   "3#冲渣泵电动阀开" AT %Q22.5 : Bool;
   "3#冲渣泵电动阀关" AT %Q22.6 : Bool;
   "3#冲渣泵排气电磁阀" AT %Q22.7 : Bool;
   "2#冲渣泵引水电磁阀" AT %Q23.0 : Bool;
   "2#冲渣泵电动阀开" AT %Q23.1 : Bool;
   "2#冲渣泵电动阀关" AT %Q23.2 : Bool;
   "2#冲渣泵排气电磁阀" AT %Q23.3 : Bool;
   "1#冲渣泵引水电磁阀" AT %Q23.4 : Bool;
   "1#冲渣泵电动阀开" AT %Q23.5 : Bool;
   "1#冲渣泵电动阀关" AT %Q23.6 : Bool;
   "1#冲渣泵排气电磁阀" AT %Q23.7 : Bool;
   "1#冲渣泵管道压力" AT %IW368 : Int;
   "2#冲渣泵管道压力" AT %IW370 : Int;
   "3#冲渣泵管道压力" AT %IW372 : Int;
   "4#冲渣泵管道压力" AT %IW374 : Int;
   "5#冲渣泵管道压力" AT %IW376 : Int;
   "6#冲渣泵管道压力" AT %IW378 : Int;
   "7#冲渣泵管道压力" AT %IW380 : Int;
   "8#冲渣泵管道压力" AT %IW382 : Int;
   "1#冲渣阀门开度" AT %IW384 : Int;
   "2#冲渣阀门开度" AT %IW386 : Int;
   "3#冲渣阀门开度" AT %IW388 : Int;
   "4#冲渣阀门开度" AT %IW390 : Int;
   "5#冲渣阀门开度" AT %IW392 : Int;
   "6#冲渣阀门开度" AT %IW394 : Int;
   "7#冲渣阀门开度" AT %IW396 : Int;
   "8#冲渣阀门开度" AT %IW398 : Int;
   "1#冲渣泵阀门开度给定" AT %QW320 : Int;
   "2#冲渣泵阀门开度给定" AT %QW322 : Int;
   "3#冲渣泵阀门开度给定" AT %QW324 : Int;
   "4#冲渣泵阀门开度给定" AT %QW326 : Int;
   "5#冲渣泵阀门开度给定" AT %QW328 : Int;
   "6#冲渣泵阀门开度给定" AT %QW330 : Int;
   "7#冲渣泵阀门开度给定" AT %QW332 : Int;
   "8#冲渣泵阀门开度给定" AT %QW334 : Int;
   "窑冷却泵运行" AT %I23.6 : Bool;
   "窑冷却泵故障" AT %I23.7 : Bool;
   "窑冷却泵驱动" AT %Q4.7 : Bool;
   "5#净环热水泵驱动" AT %Q5.0 : Bool;
   "Q5_1" AT %Q5.1 : Bool;
   "Q5_2" AT %Q5.2 : Bool;
   "Q5_3" AT %Q5.3 : Bool;
   "Q5_4" AT %Q5.4 : Bool;
   "Q5_5" AT %Q5.5 : Bool;
   "Q5_6" AT %Q5.6 : Bool;
   "Q5_7" AT %Q5.7 : Bool;
   "Q6_0" AT %Q6.0 : Bool;
   "Q6_1" AT %Q6.1 : Bool;
   "Q6_2" AT %Q6.2 : Bool;
   "Q6_3" AT %Q6.3 : Bool;
   "Q6_4" AT %Q6.4 : Bool;
   "Q6_5" AT %Q6.5 : Bool;
   "Q6_6" AT %Q6.6 : Bool;
   "Q6_7" AT %Q6.7 : Bool;
   "Q7_0" AT %Q7.0 : Bool;
   "Q7_1" AT %Q7.1 : Bool;
   "Q7_2" AT %Q7.2 : Bool;
   "Q7_3" AT %Q7.3 : Bool;
   "Q7_4" AT %Q7.4 : Bool;
   "Q7_5" AT %Q7.5 : Bool;
   "Q7_6" AT %Q7.6 : Bool;
   "Q7_7" AT %Q7.7 : Bool;
   "I32_6" AT %I32.6 : Bool;
   "I32_7" AT %I32.7 : Bool;
   "窑冷却泵电动蝶阀备妥" AT %I33.0 : Bool;
   "窑冷却泵电动蝶阀运行" AT %I33.1 : Bool;
   "窑冷却泵电动蝶阀故障" AT %I33.2 : Bool;
   "窑冷却泵电动蝶阀开到位" AT %I33.3 : Bool;
   "窑冷却泵电动蝶阀关到位" AT %I33.4 : Bool;
   "I33_5" AT %I33.5 : Bool;
   "I33_6" AT %I33.6 : Bool;
   "I33_7" AT %I33.7 : Bool;
   "I34_0" AT %I34.0 : Bool;
   "I34_1" AT %I34.1 : Bool;
   "I34_2" AT %I34.2 : Bool;
   "I34_3" AT %I34.3 : Bool;
   "I34_4" AT %I34.4 : Bool;
   "I34_5" AT %I34.5 : Bool;
   "I34_6" AT %I34.6 : Bool;
   "I34_7" AT %I34.7 : Bool;
   "I35_0" AT %I35.0 : Bool;
   "I35_1" AT %I35.1 : Bool;
   "I35_2" AT %I35.2 : Bool;
   "I35_3" AT %I35.3 : Bool;
   "I35_4" AT %I35.4 : Bool;
   "I35_5" AT %I35.5 : Bool;
   "I35_6" AT %I35.6 : Bool;
   "I35_7" AT %I35.7 : Bool;
   "5#净环热水泵电动阀开" AT %Q14.0 : Bool;
   "5#净环热水泵电动阀关" AT %Q14.1 : Bool;
   "窑冷却泵电动阀开" AT %Q14.2 : Bool;
   "窑冷却泵电动阀关" AT %Q14.3 : Bool;
   "1#柴油泵电动阀开" AT %Q14.4 : Bool;
   "1#柴油泵电动阀关" AT %Q14.5 : Bool;
   "2#柴油泵电动阀开" AT %Q14.6 : Bool;
   "2#柴油泵电动阀关" AT %Q14.7 : Bool;
   "Q15_0" AT %Q15.0 : Bool;
   "Q15_1" AT %Q15.1 : Bool;
   "Q15_2" AT %Q15.2 : Bool;
   "Q15_3" AT %Q15.3 : Bool;
   "Q15_4" AT %Q15.4 : Bool;
   "Q15_5" AT %Q15.5 : Bool;
   "Q15_6" AT %Q15.6 : Bool;
   "Q15_7" AT %Q15.7 : Bool;
   "PIW322" AT %IW322 : Int;
   "PIW324" AT %IW324 : Int;
   "PIW326" AT %IW326 : Int;
   "PIW328" AT %IW328 : Int;
   "PIW330" AT %IW330 : Int;
   "PIW332" AT %IW332 : Int;
   "PIW334" AT %IW334 : Int;
   "PQW290" AT %QW290 : Int;
   "PQW292" AT %QW292 : Int;
   "PQW294" AT %QW294 : Int;
   "PQW296" AT %QW296 : Int;
   "PQW298" AT %QW298 : Int;
   "PQW300" AT %QW300 : Int;
   "PQW302" AT %QW302 : Int;
   "I41_0" AT %I41.0 : Bool;
   "I41_1" AT %I41.1 : Bool;
   "I41_2" AT %I41.2 : Bool;
   "I41_3" AT %I41.3 : Bool;
   "I41_4" AT %I41.4 : Bool;
   "I41_5" AT %I41.5 : Bool;
   "I41_6" AT %I41.6 : Bool;
   "I41_7" AT %I41.7 : Bool;
   "I42_0" AT %I42.0 : Bool;
   "I42_1" AT %I42.1 : Bool;
   "I42_2" AT %I42.2 : Bool;
   "I42_3" AT %I42.3 : Bool;
   "I42_4" AT %I42.4 : Bool;
   "I42_5" AT %I42.5 : Bool;
   "I42_6" AT %I42.6 : Bool;
   "I42_7" AT %I42.7 : Bool;
   "I43_0" AT %I43.0 : Bool;
   "I43_1" AT %I43.1 : Bool;
   "I43_2" AT %I43.2 : Bool;
   "I43_3" AT %I43.3 : Bool;
   "I43_4" AT %I43.4 : Bool;
   "I43_5" AT %I43.5 : Bool;
   "I43_6" AT %I43.6 : Bool;
   "I43_7" AT %I43.7 : Bool;
   "I49_0" AT %I49.0 : Bool;
   "I49_1" AT %I49.1 : Bool;
   "I49_2" AT %I49.2 : Bool;
   "I49_3" AT %I49.3 : Bool;
   "I49_4" AT %I49.4 : Bool;
   "I49_5" AT %I49.5 : Bool;
   "I49_6" AT %I49.6 : Bool;
   "I49_7" AT %I49.7 : Bool;
   "I50_0" AT %I50.0 : Bool;
   "I50_1" AT %I50.1 : Bool;
   "I50_2" AT %I50.2 : Bool;
   "I50_3" AT %I50.3 : Bool;
   "I50_4" AT %I50.4 : Bool;
   "I50_5" AT %I50.5 : Bool;
   "I50_6" AT %I50.6 : Bool;
   "I50_7" AT %I50.7 : Bool;
   "I51_0" AT %I51.0 : Bool;
   "I51_1" AT %I51.1 : Bool;
   "I51_2" AT %I51.2 : Bool;
   "I51_3" AT %I51.3 : Bool;
   "I51_4" AT %I51.4 : Bool;
   "I51_5" AT %I51.5 : Bool;
   "I51_6" AT %I51.6 : Bool;
   "I51_7" AT %I51.7 : Bool;
   "Tag_1" AT %M1.4 : Bool;
   "Tag_2" AT %M2.0 : Bool;
   "Tag_3" AT %T40 : Timer;
   "Tag_4" AT %M2.1 : Bool;
   "Tag_5" AT %MW4 : Int;
   "Tag_6" AT %M2.2 : Bool;
   "Tag_7" AT %M2.3 : Bool;
   "Tag_8" AT %M2.4 : Bool;
   "Tag_9" AT %M2.5 : Bool;
   "Tag_10" AT %M2.6 : Bool;
   "Tag_11" AT %M2.7 : Bool;
   "Tag_12" AT %M3.0 : Bool;
   "Tag_13" AT %M3.1 : Bool;
   "Tag_14" AT %M3.2 : Bool;
   "Tag_15" AT %MD4 : Real;
   "Tag_16" AT %MD8 : Real;
   "HMI_允许电炉启动冲渣泵1" AT %M100.0 : Bool;
   "HMI_允许电炉启动冲渣泵2" AT %M100.1 : Bool;
   "HMI_允许电炉启动冲渣泵3" AT %M100.2 : Bool;
   "HMI_允许电炉启动冲渣泵4" AT %M100.3 : Bool;
   "HMI_允许电炉启动冲渣泵5" AT %M100.4 : Bool;
   "HMI_允许电炉启动冲渣泵6" AT %M100.5 : Bool;
   "HMI_允许电炉启动冲渣泵7" AT %M100.6 : Bool;
   "HMI_允许电炉启动冲渣泵8" AT %M100.7 : Bool;
   "HMI_电炉冲渣急停1" AT %M99.0 : Bool;
   "HMI_电炉冲渣急停2" AT %M99.1 : Bool;
   "Tag_17" AT %M11.1 : Bool;
END_VAR

DATA_BLOCK "AI"   // DB2
{ S7_Optimized_Access := 'FALSE' }
VERSION : 0.1
   VAR
      "1#炉体水泵管道压力" : Real;
      "2#炉体水泵管道压力" : Real;
      "3#炉体水泵管道压力" : Real;
      "1#电极水泵管道压力" : Real;
      "2#电极水泵管道压力" : Real;
      "3#电极水泵管道压力" : Real;
      "4#电极水泵管道压力" : Real;
      "1#柴油泵管道压力" : Real;
      "2#柴油泵管道压力" : Real;
      "1#炉体水阀门开度" : Real;
      "2#炉体水阀门开度" : Real;
      "3#炉体水阀门开度" : Real;
      "1#电极水阀门开度" : Real;
      "2#电极水阀门开度" : Real;
      "3#电极水阀门开度" : Real;
      "4#电极水阀门开度" : Real;
      "2#柴油泵阀门开度" : Real;
      "1#净环热水管道压力" : Real;
      "2#净环热水管道压力" : Real;
      "3#净环热水管道压力" : Real;
      "4#净环热水管道压力" : Real;
      "5#净环热水管道压力" : Real;
      "6#净环热水管道压力" : Real;
      "1#净环热水阀门开度" : Real;
      "2#净环热水阀门开度" : Real;
      "3#净环热水阀门开度" : Real;
      "4#净环热水阀门开度" : Real;
      "5#净环热水阀门开度" : Real;
      "6#净环热水阀门开度" : Real;
      "1#外围补水阀门开度" : Real;
      "2#外围补水阀门开度" : Real;
      "1#水池液位" : Real;
      "2#水池液位" : Real;
      PIW322 : Real;
      PIW324 : Real;
      PIW326 : Real;
      PIW328 : Real;
      PIW330 : Real;
      PIW332 : Real;
      PIW334 : Real;
      "1#冲渣热水泵管道压力" : Real;
      "2#冲渣热水泵管道压力" : Real;
      "3#冲渣热水泵管道压力" : Real;
      "4#冲渣热水泵管道压力" : Real;
      "5#冲渣热水泵管道压力" : Real;
      "6#冲渣热水泵管道压力" : Real;
      "7#冲渣热水泵管道压力" : Real;
      "8#冲渣热水泵管道压力" : Real;
      "1#冲渣热水阀门开度" : Real;
      "2#冲渣热水阀门开度" : Real;
      "3#冲渣热水阀门开度" : Real;
      "4#冲渣热水阀门开度" : Real;
      "5#冲渣热水阀门开度" : Real;
      "6#冲渣热水阀门开度" : Real;
      "7#冲渣热水阀门开度" : Real;
      "8#冲渣热水阀门开度" : Real;
      "1#冲渣泵管道压力" : Real;
      "2#冲渣泵管道压力" : Real;
      "3#冲渣泵管道压力" : Real;
      "4#冲渣泵管道压力" : Real;
      "5#冲渣泵管道压力" : Real;
      "6#冲渣泵管道压力" : Real;
      "7#冲渣泵管道压力" : Real;
      "8#冲渣泵管道压力" : Real;
      "1#冲渣阀门开度" : Real;
      "2#冲渣阀门开度" : Real;
      "3#冲渣阀门开度" : Real;
      "4#冲渣阀门开度" : Real;
      "5#冲渣阀门开度" : Real;
      "6#冲渣阀门开度" : Real;
      "7#冲渣阀门开度" : Real;
      "8#冲渣阀门开度" : Real;
      Static1 : Real;
      Static2 : Real;
      Static3 : Real;
      Static4 : Real;
      Static5 : Real;
      Static6 : Real;
      Static7 : Real;
      Static8 : Real;
      Static9 : Real;
      Static10 : Real;
      Static11 : Real;
      Static12 : Real;
      Static13 : Real;
      Static14 : Real;
      Static15 : Real;
      Static16 : Real;
      Static17 : Real;
      Static18 : Real;
      Static19 : Real;
      Static20 : Real;
      Static21 : Real;
      Static22 : Real;
      Static23 : Real;
      Static24 : Real;
      Static25 : Real;
      Static26 : Real;
      Static27 : Real;
      Static28 : Real;
      Static29 : Real;
      Static30 : Real;
      Static31 : Real;
      Static32 : Real;
      Static33 : Real;
      Static34 : Real;
      Static35 : Real;
      Static36 : Real;
      Static37 : Real;
      Static38 : Real;
      Static39 : Real;
      Static40 : Real;
      Static41 : Real;
      Static42 : Real;
      Static43 : Real;
      Static44 : Real;
      Static45 : Real;
      Static46 : Real;
      Static47 : Real;
      Static48 : Real;
      Static49 : Real;
      Static50 : Real;
      Static51 : Real;
      Static52 : Real;
      Static53 : Real;
      Static54 : Real;
      Static55 : Real;
      Static56 : Real;
      Static57 : Real;
      Static58 : Real;
      Static59 : Real;
      Static60 : Real;
      Static61 : Real;
      Static62 : Real;
      Static63 : Real;
      Static64 : Real;
      Static65 : Real;
      Static66 : Real;
      Static67 : Real;
      Static68 : Real;
      Static69 : Real;
      Static70 : Real;
      Static71 : Real;
      Static72 : Real;
      Static73 : Real;
      Static74 : Real;
      Static75 : Real;
      Static76 : Real;
      Static77 : Real;
      Static78 : Real;
      Static79 : Real;
      Static80 : Real;
      Static81 : Real;
      Static82 : Real;
      Static83 : Real;
      Static84 : Real;
      Static85 : Real;
      Static86 : Real;
      Static87 : Real;
      Static88 : Real;
      Static89 : Real;
      Static90 : Real;
      Static91 : Real;
      Static92 : Real;
      Static93 : Real;
      Static94 : Real;
      Static95 : Real;
      Static96 : Real;
      Static97 : Real;
      Static98 : Real;
      Static99 : Real;
   END_VAR
BEGIN
END_DATA_BLOCK

DATA_BLOCK "AO"   // DB3
{ S7_Optimized_Access := 'TRUE' }
VERSION : 0.1
   VAR
      "1#循环水泵阀门开度给定" : Real := 0.0;
      "2#循环水泵阀门开度给定" : Real := 0.0;
      "3#循环水泵阀门开度给定" : Real := 0.0;
      "1#电极冷却泵阀门开度给定" : Real := 0.0;
      "2#电极冷却泵阀门开度给定" : Real := 0.0;
      "3#电极冷却泵阀门开度给定" : Real := 0.0;
      "4#电极冷却泵阀门开度给定" : Real := 0.0;
      "1#柴油泵阀门开度给定" : Real := 0.0;
      "2#柴油泵阀门开度给定" : Real := 0.0;
      "1#净环热水泵阀门开度给定" : Real := 0.0;
      "2#净环热水泵阀门开度给定" : Real := 0.0;
      "3#净环热水泵阀门开度给定" : Real := 0.0;
      "4#净环热水泵阀门开度给定" : Real := 0.0;
      "5#净环热水泵阀门开度给定" : Real := 0.0;
      "6#净环热水泵阀门开度给定" : Real := 0.0;
      "1#外围补水阀门开度给定" : Real := 0.0;
      "2#外围补水阀门开度给定" : Real := 0.0;
      PQW290 : Real := 0.0;   // useless
      PQW292 : Real := 0.0;
      PQW294 : Real := 0.0;
      PQW296 : Real := 0.0;
      PQW298 : Real := 0.0;
      PQW300 : Real := 0.0;
      PQW302 : Real := 0.0;
      "1#冲渣热水泵阀门开度给定" : Real := 0.0;
      "2#冲渣热水泵阀门开度给定" : Real := 0.0;
      "3#冲渣热水泵阀门开度给定" : Real := 0.0;
      "4#冲渣热水泵阀门开度给定" : Real := 0.0;
      "5#冲渣热水泵阀门开度给定" : Real := 0.0;
      "6#冲渣热水泵阀门开度给定" : Real := 0.0;
      "7#冲渣热水泵阀门开度给定" : Real := 0.0;
      "8#冲渣热水泵阀门开度给定" : Real := 0.0;
      "1#冲渣泵阀门开度给定" : Real := 0.0;
      "2#冲渣泵阀门开度给定" : Real := 0.0;
      "3#冲渣泵阀门开度给定" : Real := 0.0;
      "4#冲渣泵阀门开度给定" : Real := 0.0;
      "5#冲渣泵阀门开度给定" : Real := 0.0;
      "6#冲渣泵阀门开度给定" : Real := 0.0;
      "7#冲渣泵阀门开度给定" : Real := 0.0;
      "8#冲渣泵阀门开度给定" : Real := 0.0;
      Static1 : Real := 0.0;
      Static2 : Real := 0.0;
      Static3 : Real := 0.0;
      Static4 : Real := 0.0;
      Static5 : Real := 0.0;
      Static6 : Real := 0.0;
      Static7 : Real := 0.0;
      Static8 : Real := 0.0;
      Static9 : Real := 0.0;
      Static10 : Real := 0.0;
      Static11 : Real := 0.0;
      Static12 : Real := 0.0;
      Static13 : Real := 0.0;
      Static14 : Real := 0.0;
      Static15 : Real := 0.0;
      Static16 : Real := 0.0;
      Static17 : Real := 0.0;
      Static18 : Real := 0.0;
      Static19 : Real := 0.0;
      Static20 : Real := 0.0;
      Static21 : Real := 0.0;
      Static22 : Real := 0.0;
      Static23 : Real := 0.0;
      Static24 : Real := 0.0;
      Static25 : Real := 0.0;
      Static26 : Real := 0.0;
      Static27 : Real := 0.0;
      Static28 : Real := 0.0;
      Static29 : Real := 0.0;
      Static30 : Real := 0.0;
      Static31 : Real := 0.0;
      Static32 : Real := 0.0;
      Static33 : Real := 0.0;
      Static34 : Real := 0.0;
      Static35 : Real := 0.0;
      Static36 : Real := 0.0;
      Static37 : Real := 0.0;
      Static38 : Real := 0.0;
      Static39 : Real := 0.0;
      Static40 : Real := 0.0;
      Static41 : Real := 0.0;
      Static42 : Real := 0.0;
      Static43 : Real := 0.0;
      Static44 : Real := 0.0;
      Static45 : Real := 0.0;
      Static46 : Real := 0.0;
      Static47 : Real := 0.0;
      Static48 : Real := 0.0;
      Static49 : Real := 0.0;
      Static50 : Real := 0.0;
      Static51 : Real := 0.0;
      Static52 : Real := 0.0;
      Static53 : Real := 0.0;
      Static54 : Real := 0.0;
      Static55 : Real := 0.0;
      Static56 : Real := 0.0;
      Static57 : Real := 0.0;
      Static58 : Real := 0.0;
      Static99 : Real := 0.0;
   END_VAR
BEGIN
END_DATA_BLOCK

DATA_BLOCK "TIME"   // DB4
{ S7_Optimized_Access := 'TRUE' }
VERSION : 0.1
   VAR
      T1 : IEC_TIMER;
      T2 : IEC_TIMER;
      T3 : IEC_TIMER;
      T4 : IEC_TIMER;
      T5 : IEC_TIMER;
      T6 : IEC_TIMER;
      T7 : IEC_TIMER;
      T8 : IEC_TIMER;
      T9 : IEC_TIMER;
      T10 : IEC_TIMER;
      T11 : IEC_TIMER;
      T12 : IEC_TIMER;
      T13 : IEC_TIMER;
      T14 : IEC_TIMER;
      T15 : IEC_TIMER;
      T16 : IEC_TIMER;
      T17 : IEC_TIMER;
      T18 : IEC_TIMER;
      T19 : IEC_TIMER;
      T20 : IEC_TIMER;
      T21 : IEC_TIMER;
      T22 : IEC_TIMER;
      T23 : IEC_TIMER;
      T24 : IEC_TIMER;
      T25 : IEC_TIMER;
      T26 : IEC_TIMER;
      T27 : IEC_TIMER;
      T28 : IEC_TIMER;
   END_VAR
BEGIN
END_DATA_BLOCK

DATA_BLOCK "DB15_PLC_TO_HMI"   // DB5
{ S7_Optimized_Access := 'FALSE' }
VERSION : 0.1
   VAR
      P1 : Bool;
      P2 : Bool;
      P3 : Bool;
      P4 : Bool;
      P5 : Bool;
      P6 : Bool;
      P7 : Bool;
      P8 : Bool;
      P9 : Bool;
      P10 : Bool;
      P11 : Bool;
      P12 : Bool;
      P13 : Bool;
      P14 : Bool;
      P15 : Bool;
      P16 : Bool;
      HMI_电炉冲渣急停1次数 : Int;
      HMI_电炉冲渣急停2次数 : Int;
      static1 : Int;
      static2 : Int;
      static3 : Int;
      static4 : Int;
      static5 : Int;
      static6 : Int;
      static7 : Int;
      static8 : Int;
      static9 : Int;
      static10 : Int;
      static11 : Int;
      static12 : Int;
   END_VAR
BEGIN
END_DATA_BLOCK

DATA_BLOCK "电机_冷却塔风机FB_DB"   // DB10
{ S7_Optimized_Access := 'FALSE' }
VERSION : 0.1
// stored: InstanceOfName 电机_冷却塔风机FB
"电机_冷却塔风机FB"
BEGIN
END_DATA_BLOCK

DATA_BLOCK "阀门_FB_DB"   // DB11
{ S7_Optimized_Access := 'FALSE' }
VERSION : 0.1
// stored: InstanceOfName 阀门_FB
"阀门_FB"
BEGIN
END_DATA_BLOCK

DATA_BLOCK "引水阀和排气阀FB_DB"   // DB12
{ S7_Optimized_Access := 'FALSE' }
VERSION : 0.1
// stored: InstanceOfName 引水阀和排气阀FB
"引水阀和排气阀FB"
BEGIN
END_DATA_BLOCK

DATA_BLOCK "电机_泵FB_DB"   // DB13
{ S7_Optimized_Access := 'FALSE' }
VERSION : 0.1
// stored: InstanceOfName 电机_泵FB
"电机_泵FB"
BEGIN
END_DATA_BLOCK

DATA_BLOCK "FB14_DATA_ALARM_DB"   // DB14
{ S7_Optimized_Access := 'FALSE' }
VERSION : 0.1
// stored: InstanceOfName FB14_DATA_ALARM
"FB14_DATA_ALARM"
BEGIN
END_DATA_BLOCK

DATA_BLOCK "FB15_MOTOR_AUTO-st_DB"   // DB15
{ S7_Optimized_Access := 'FALSE' }
VERSION : 0.1
// stored: InstanceOfName FB15_MOTOR_AUTO-st
"FB15_MOTOR_AUTO-st"
BEGIN
END_DATA_BLOCK

FUNCTION_BLOCK "电机_冷却塔风机FB"   // FB10, LAD
{ S7_Optimized_Access := 'FALSE' }
VERSION : 0.1
   VAR
      "1#冲渣水池冷却塔风机" : "电机_冷却塔风机";
      "2#冲渣水池冷却塔风机" : "电机_冷却塔风机";
      "3#冲渣水池冷却塔风机" : "电机_冷却塔风机";
      "4#冲渣水池冷却塔风机" : "电机_冷却塔风机";
      "5#冲渣水池冷却塔风机" : "电机_冷却塔风机";
      "6#冲渣水池冷却塔风机" : "电机_冷却塔风机";
      "1#净环水池冷却塔风机" : "电机_冷却塔风机";
      "2#净环水池冷却塔风机" : "电机_冷却塔风机";
      "3#净环水池冷却塔风机" : "电机_冷却塔风机";
      "4#净环水池冷却塔风机" : "电机_冷却塔风机";
      备用1 : "电机_冷却塔风机";
      备用2 : "电机_冷却塔风机";
      备用3 : "电机_冷却塔风机";
      备用4 : "电机_冷却塔风机";
      备用5 : "电机_冷却塔风机";
      备用6 : "电机_冷却塔风机";
      备用7 : "电机_冷却塔风机";
      备用8 : "电机_冷却塔风机";
      备用9 : "电机_冷却塔风机";
      备用10 : "电机_冷却塔风机";
   END_VAR
BEGIN

REGION Network 1
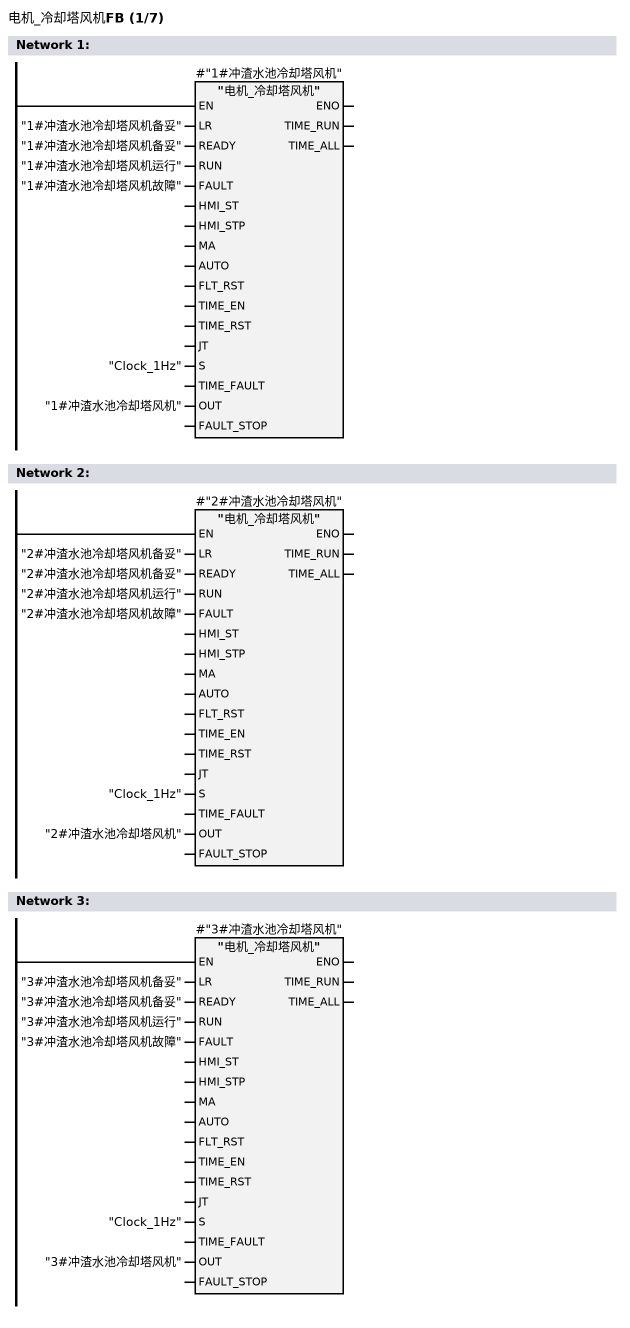
   RUNG wire#powerrail
      #"1#冲渣水池冷却塔风机"(LR := "1#冲渣水池冷却塔风机备妥", READY := "1#冲渣水池冷却塔风机备妥", RUN := "1#冲渣水池冷却塔风机运行", FAULT := "1#冲渣水池冷却塔风机故障", HMI_ST :=, HMI_STP :=, MA :=, AUTO :=, FLT_RST :=, TIME_EN :=, TIME_RST :=, JT :=, S := "Clock_1Hz", TIME_FAULT :=, OUT := "1#冲渣水池冷却塔风机", FAULT_STOP :=, TIME_RUN =>, TIME_ALL =>)
   END_RUNG
   // the same network as SCL:
   #"1#冲渣水池冷却塔风机"(LR := "1#冲渣水池冷却塔风机备妥",   // "电机_冷却塔风机"
                  READY := "1#冲渣水池冷却塔风机备妥",
                  RUN := "1#冲渣水池冷却塔风机运行",
                  FAULT := "1#冲渣水池冷却塔风机故障",
                  S := "Clock_1Hz",
                  OUT := "1#冲渣水池冷却塔风机");
END_REGION

REGION Network 2
   RUNG wire#powerrail
      #"2#冲渣水池冷却塔风机"(LR := "2#冲渣水池冷却塔风机备妥", READY := "2#冲渣水池冷却塔风机备妥", RUN := "2#冲渣水池冷却塔风机运行", FAULT := "2#冲渣水池冷却塔风机故障", HMI_ST :=, HMI_STP :=, MA :=, AUTO :=, FLT_RST :=, TIME_EN :=, TIME_RST :=, JT :=, S := "Clock_1Hz", TIME_FAULT :=, OUT := "2#冲渣水池冷却塔风机", FAULT_STOP :=, TIME_RUN =>, TIME_ALL =>)
   END_RUNG
   // the same network as SCL:
   #"2#冲渣水池冷却塔风机"(LR := "2#冲渣水池冷却塔风机备妥",   // "电机_冷却塔风机"
                  READY := "2#冲渣水池冷却塔风机备妥",
                  RUN := "2#冲渣水池冷却塔风机运行",
                  FAULT := "2#冲渣水池冷却塔风机故障",
                  S := "Clock_1Hz",
                  OUT := "2#冲渣水池冷却塔风机");
END_REGION

REGION Network 3
   RUNG wire#powerrail
      #"3#冲渣水池冷却塔风机"(LR := "3#冲渣水池冷却塔风机备妥", READY := "3#冲渣水池冷却塔风机备妥", RUN := "3#冲渣水池冷却塔风机运行", FAULT := "3#冲渣水池冷却塔风机故障", HMI_ST :=, HMI_STP :=, MA :=, AUTO :=, FLT_RST :=, TIME_EN :=, TIME_RST :=, JT :=, S := "Clock_1Hz", TIME_FAULT :=, OUT := "3#冲渣水池冷却塔风机", FAULT_STOP :=, TIME_RUN =>, TIME_ALL =>)
   END_RUNG
   // the same network as SCL:
   #"3#冲渣水池冷却塔风机"(LR := "3#冲渣水池冷却塔风机备妥",   // "电机_冷却塔风机"
                  READY := "3#冲渣水池冷却塔风机备妥",
                  RUN := "3#冲渣水池冷却塔风机运行",
                  FAULT := "3#冲渣水池冷却塔风机故障",
                  S := "Clock_1Hz",
                  OUT := "3#冲渣水池冷却塔风机");
END_REGION

REGION Network 4
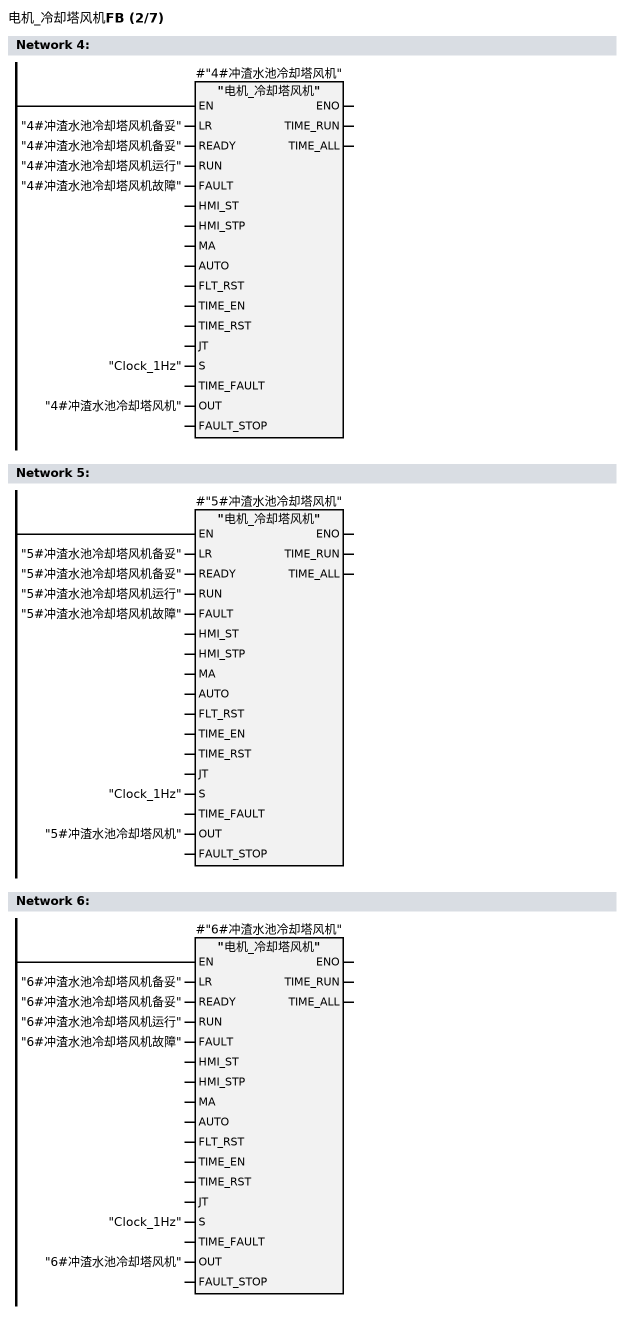
   RUNG wire#powerrail
      #"4#冲渣水池冷却塔风机"(LR := "4#冲渣水池冷却塔风机备妥", READY := "4#冲渣水池冷却塔风机备妥", RUN := "4#冲渣水池冷却塔风机运行", FAULT := "4#冲渣水池冷却塔风机故障", HMI_ST :=, HMI_STP :=, MA :=, AUTO :=, FLT_RST :=, TIME_EN :=, TIME_RST :=, JT :=, S := "Clock_1Hz", TIME_FAULT :=, OUT := "4#冲渣水池冷却塔风机", FAULT_STOP :=, TIME_RUN =>, TIME_ALL =>)
   END_RUNG
   // the same network as SCL:
   #"4#冲渣水池冷却塔风机"(LR := "4#冲渣水池冷却塔风机备妥",   // "电机_冷却塔风机"
                  READY := "4#冲渣水池冷却塔风机备妥",
                  RUN := "4#冲渣水池冷却塔风机运行",
                  FAULT := "4#冲渣水池冷却塔风机故障",
                  S := "Clock_1Hz",
                  OUT := "4#冲渣水池冷却塔风机");
END_REGION

REGION Network 5
   RUNG wire#powerrail
      #"5#冲渣水池冷却塔风机"(LR := "5#冲渣水池冷却塔风机备妥", READY := "5#冲渣水池冷却塔风机备妥", RUN := "5#冲渣水池冷却塔风机运行", FAULT := "5#冲渣水池冷却塔风机故障", HMI_ST :=, HMI_STP :=, MA :=, AUTO :=, FLT_RST :=, TIME_EN :=, TIME_RST :=, JT :=, S := "Clock_1Hz", TIME_FAULT :=, OUT := "5#冲渣水池冷却塔风机", FAULT_STOP :=, TIME_RUN =>, TIME_ALL =>)
   END_RUNG
   // the same network as SCL:
   #"5#冲渣水池冷却塔风机"(LR := "5#冲渣水池冷却塔风机备妥",   // "电机_冷却塔风机"
                  READY := "5#冲渣水池冷却塔风机备妥",
                  RUN := "5#冲渣水池冷却塔风机运行",
                  FAULT := "5#冲渣水池冷却塔风机故障",
                  S := "Clock_1Hz",
                  OUT := "5#冲渣水池冷却塔风机");
END_REGION

REGION Network 6
   RUNG wire#powerrail
      #"6#冲渣水池冷却塔风机"(LR := "6#冲渣水池冷却塔风机备妥", READY := "6#冲渣水池冷却塔风机备妥", RUN := "6#冲渣水池冷却塔风机运行", FAULT := "6#冲渣水池冷却塔风机故障", HMI_ST :=, HMI_STP :=, MA :=, AUTO :=, FLT_RST :=, TIME_EN :=, TIME_RST :=, JT :=, S := "Clock_1Hz", TIME_FAULT :=, OUT := "6#冲渣水池冷却塔风机", FAULT_STOP :=, TIME_RUN =>, TIME_ALL =>)
   END_RUNG
   // the same network as SCL:
   #"6#冲渣水池冷却塔风机"(LR := "6#冲渣水池冷却塔风机备妥",   // "电机_冷却塔风机"
                  READY := "6#冲渣水池冷却塔风机备妥",
                  RUN := "6#冲渣水池冷却塔风机运行",
                  FAULT := "6#冲渣水池冷却塔风机故障",
                  S := "Clock_1Hz",
                  OUT := "6#冲渣水池冷却塔风机");
END_REGION

REGION Network 7
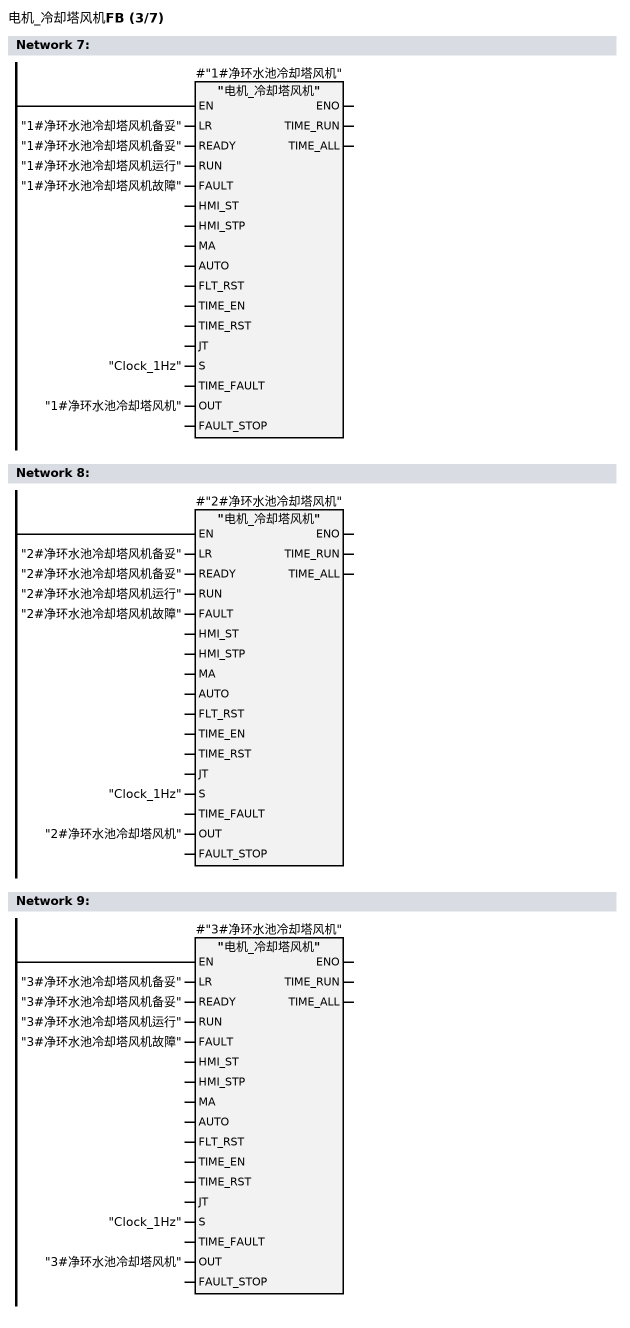
   RUNG wire#powerrail
      #"1#净环水池冷却塔风机"(LR := "1#净环水池冷却塔风机备妥", READY := "1#净环水池冷却塔风机备妥", RUN := "1#净环水池冷却塔风机运行", FAULT := "1#净环水池冷却塔风机故障", HMI_ST :=, HMI_STP :=, MA :=, AUTO :=, FLT_RST :=, TIME_EN :=, TIME_RST :=, JT :=, S := "Clock_1Hz", TIME_FAULT :=, OUT := "1#净环水池冷却塔风机", FAULT_STOP :=, TIME_RUN =>, TIME_ALL =>)
   END_RUNG
   // the same network as SCL:
   #"1#净环水池冷却塔风机"(LR := "1#净环水池冷却塔风机备妥",   // "电机_冷却塔风机"
                  READY := "1#净环水池冷却塔风机备妥",
                  RUN := "1#净环水池冷却塔风机运行",
                  FAULT := "1#净环水池冷却塔风机故障",
                  S := "Clock_1Hz",
                  OUT := "1#净环水池冷却塔风机");
END_REGION

REGION Network 8
   RUNG wire#powerrail
      #"2#净环水池冷却塔风机"(LR := "2#净环水池冷却塔风机备妥", READY := "2#净环水池冷却塔风机备妥", RUN := "2#净环水池冷却塔风机运行", FAULT := "2#净环水池冷却塔风机故障", HMI_ST :=, HMI_STP :=, MA :=, AUTO :=, FLT_RST :=, TIME_EN :=, TIME_RST :=, JT :=, S := "Clock_1Hz", TIME_FAULT :=, OUT := "2#净环水池冷却塔风机", FAULT_STOP :=, TIME_RUN =>, TIME_ALL =>)
   END_RUNG
   // the same network as SCL:
   #"2#净环水池冷却塔风机"(LR := "2#净环水池冷却塔风机备妥",   // "电机_冷却塔风机"
                  READY := "2#净环水池冷却塔风机备妥",
                  RUN := "2#净环水池冷却塔风机运行",
                  FAULT := "2#净环水池冷却塔风机故障",
                  S := "Clock_1Hz",
                  OUT := "2#净环水池冷却塔风机");
END_REGION

REGION Network 9
   RUNG wire#powerrail
      #"3#净环水池冷却塔风机"(LR := "3#净环水池冷却塔风机备妥", READY := "3#净环水池冷却塔风机备妥", RUN := "3#净环水池冷却塔风机运行", FAULT := "3#净环水池冷却塔风机故障", HMI_ST :=, HMI_STP :=, MA :=, AUTO :=, FLT_RST :=, TIME_EN :=, TIME_RST :=, JT :=, S := "Clock_1Hz", TIME_FAULT :=, OUT := "3#净环水池冷却塔风机", FAULT_STOP :=, TIME_RUN =>, TIME_ALL =>)
   END_RUNG
   // the same network as SCL:
   #"3#净环水池冷却塔风机"(LR := "3#净环水池冷却塔风机备妥",   // "电机_冷却塔风机"
                  READY := "3#净环水池冷却塔风机备妥",
                  RUN := "3#净环水池冷却塔风机运行",
                  FAULT := "3#净环水池冷却塔风机故障",
                  S := "Clock_1Hz",
                  OUT := "3#净环水池冷却塔风机");
END_REGION

REGION Network 10
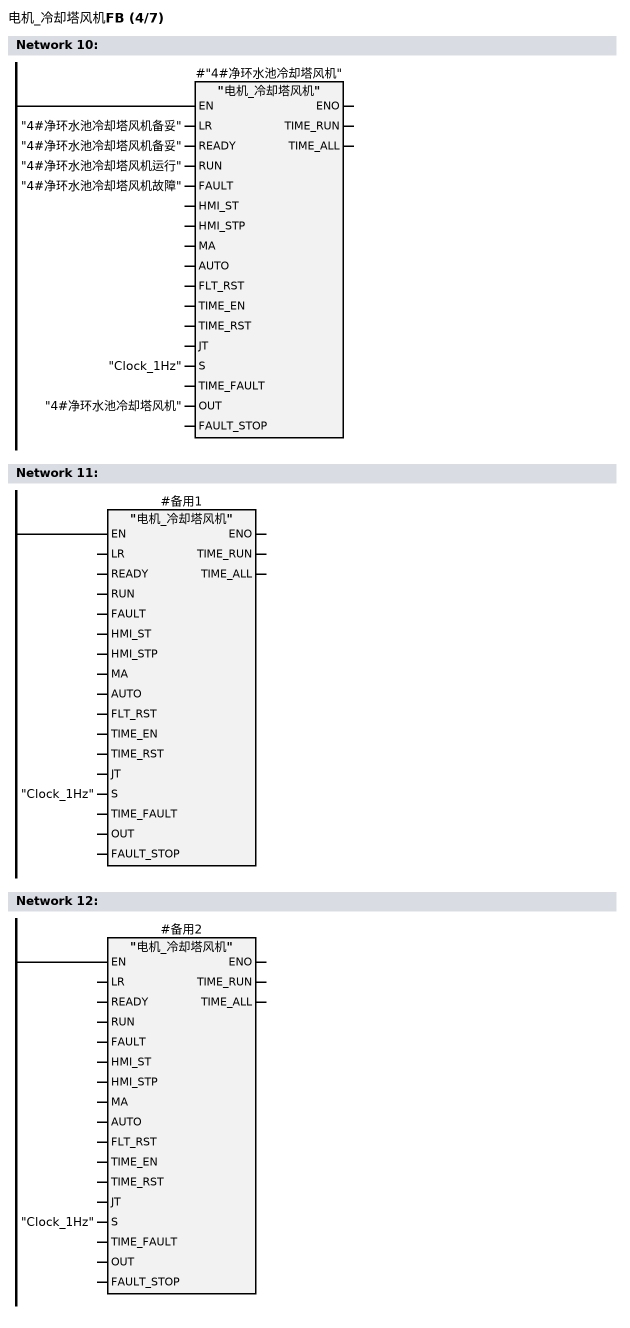
   RUNG wire#powerrail
      #"4#净环水池冷却塔风机"(LR := "4#净环水池冷却塔风机备妥", READY := "4#净环水池冷却塔风机备妥", RUN := "4#净环水池冷却塔风机运行", FAULT := "4#净环水池冷却塔风机故障", HMI_ST :=, HMI_STP :=, MA :=, AUTO :=, FLT_RST :=, TIME_EN :=, TIME_RST :=, JT :=, S := "Clock_1Hz", TIME_FAULT :=, OUT := "4#净环水池冷却塔风机", FAULT_STOP :=, TIME_RUN =>, TIME_ALL =>)
   END_RUNG
   // the same network as SCL:
   #"4#净环水池冷却塔风机"(LR := "4#净环水池冷却塔风机备妥",   // "电机_冷却塔风机"
                  READY := "4#净环水池冷却塔风机备妥",
                  RUN := "4#净环水池冷却塔风机运行",
                  FAULT := "4#净环水池冷却塔风机故障",
                  S := "Clock_1Hz",
                  OUT := "4#净环水池冷却塔风机");
END_REGION

REGION Network 11
   RUNG wire#powerrail
      #备用1(LR :=, READY :=, RUN :=, FAULT :=, HMI_ST :=, HMI_STP :=, MA :=, AUTO :=, FLT_RST :=, TIME_EN :=, TIME_RST :=, JT :=, S := "Clock_1Hz", TIME_FAULT :=, OUT :=, FAULT_STOP :=, TIME_RUN =>, TIME_ALL =>)
   END_RUNG
   // the same network as SCL:
   #备用1(S := "Clock_1Hz");   // "电机_冷却塔风机"
END_REGION

REGION Network 12
   RUNG wire#powerrail
      #备用2(LR :=, READY :=, RUN :=, FAULT :=, HMI_ST :=, HMI_STP :=, MA :=, AUTO :=, FLT_RST :=, TIME_EN :=, TIME_RST :=, JT :=, S := "Clock_1Hz", TIME_FAULT :=, OUT :=, FAULT_STOP :=, TIME_RUN =>, TIME_ALL =>)
   END_RUNG
   // the same network as SCL:
   #备用2(S := "Clock_1Hz");   // "电机_冷却塔风机"
END_REGION

REGION Network 13
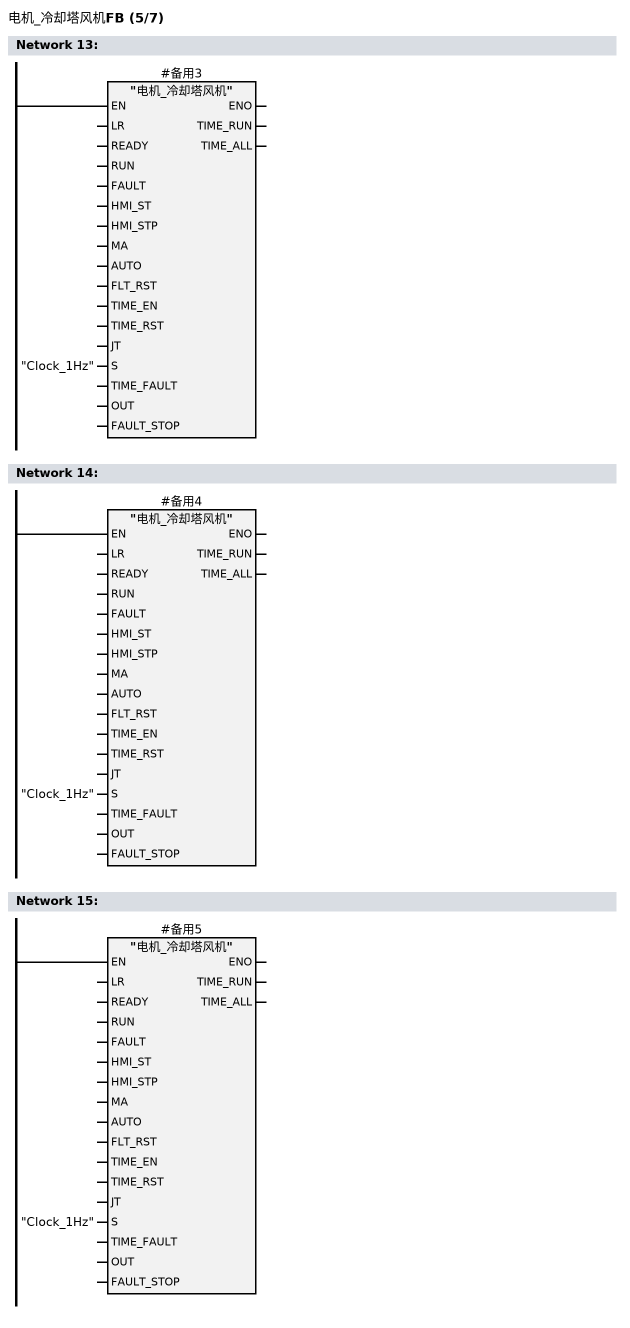
   RUNG wire#powerrail
      #备用3(LR :=, READY :=, RUN :=, FAULT :=, HMI_ST :=, HMI_STP :=, MA :=, AUTO :=, FLT_RST :=, TIME_EN :=, TIME_RST :=, JT :=, S := "Clock_1Hz", TIME_FAULT :=, OUT :=, FAULT_STOP :=, TIME_RUN =>, TIME_ALL =>)
   END_RUNG
   // the same network as SCL:
   #备用3(S := "Clock_1Hz");   // "电机_冷却塔风机"
END_REGION

REGION Network 14
   RUNG wire#powerrail
      #备用4(LR :=, READY :=, RUN :=, FAULT :=, HMI_ST :=, HMI_STP :=, MA :=, AUTO :=, FLT_RST :=, TIME_EN :=, TIME_RST :=, JT :=, S := "Clock_1Hz", TIME_FAULT :=, OUT :=, FAULT_STOP :=, TIME_RUN =>, TIME_ALL =>)
   END_RUNG
   // the same network as SCL:
   #备用4(S := "Clock_1Hz");   // "电机_冷却塔风机"
END_REGION

REGION Network 15
   RUNG wire#powerrail
      #备用5(LR :=, READY :=, RUN :=, FAULT :=, HMI_ST :=, HMI_STP :=, MA :=, AUTO :=, FLT_RST :=, TIME_EN :=, TIME_RST :=, JT :=, S := "Clock_1Hz", TIME_FAULT :=, OUT :=, FAULT_STOP :=, TIME_RUN =>, TIME_ALL =>)
   END_RUNG
   // the same network as SCL:
   #备用5(S := "Clock_1Hz");   // "电机_冷却塔风机"
END_REGION

REGION Network 16
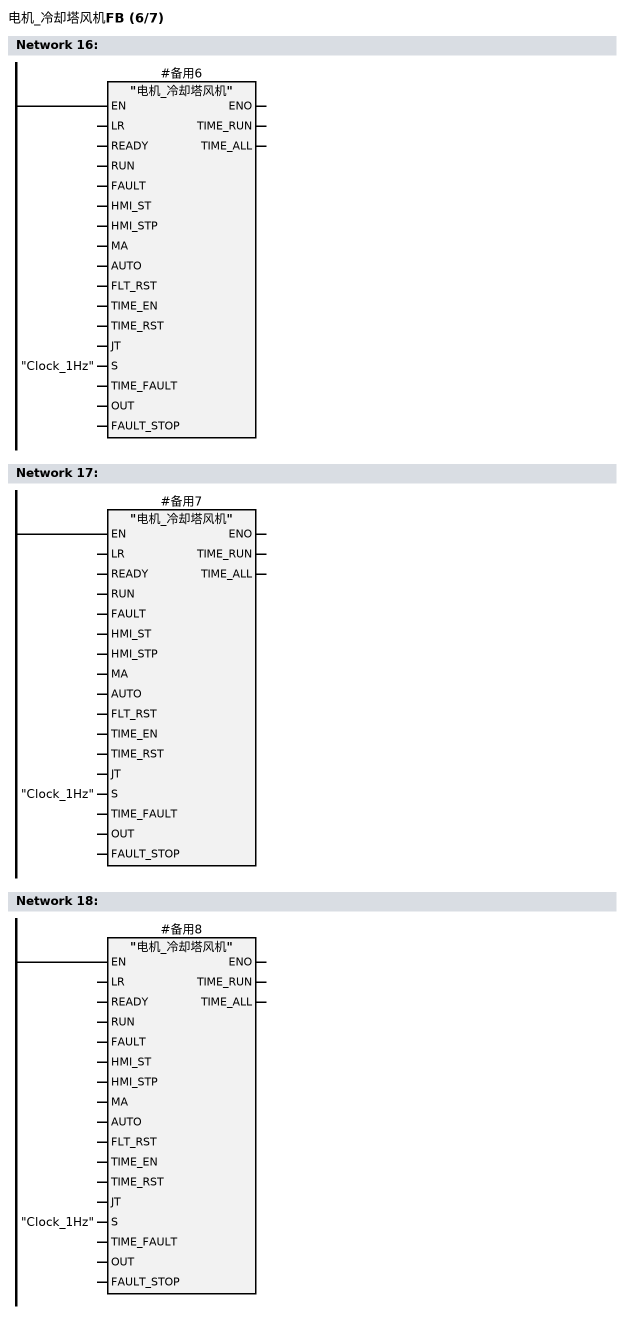
   RUNG wire#powerrail
      #备用6(LR :=, READY :=, RUN :=, FAULT :=, HMI_ST :=, HMI_STP :=, MA :=, AUTO :=, FLT_RST :=, TIME_EN :=, TIME_RST :=, JT :=, S := "Clock_1Hz", TIME_FAULT :=, OUT :=, FAULT_STOP :=, TIME_RUN =>, TIME_ALL =>)
   END_RUNG
   // the same network as SCL:
   #备用6(S := "Clock_1Hz");   // "电机_冷却塔风机"
END_REGION

REGION Network 17
   RUNG wire#powerrail
      #备用7(LR :=, READY :=, RUN :=, FAULT :=, HMI_ST :=, HMI_STP :=, MA :=, AUTO :=, FLT_RST :=, TIME_EN :=, TIME_RST :=, JT :=, S := "Clock_1Hz", TIME_FAULT :=, OUT :=, FAULT_STOP :=, TIME_RUN =>, TIME_ALL =>)
   END_RUNG
   // the same network as SCL:
   #备用7(S := "Clock_1Hz");   // "电机_冷却塔风机"
END_REGION

REGION Network 18
   RUNG wire#powerrail
      #备用8(LR :=, READY :=, RUN :=, FAULT :=, HMI_ST :=, HMI_STP :=, MA :=, AUTO :=, FLT_RST :=, TIME_EN :=, TIME_RST :=, JT :=, S := "Clock_1Hz", TIME_FAULT :=, OUT :=, FAULT_STOP :=, TIME_RUN =>, TIME_ALL =>)
   END_RUNG
   // the same network as SCL:
   #备用8(S := "Clock_1Hz");   // "电机_冷却塔风机"
END_REGION

REGION Network 19
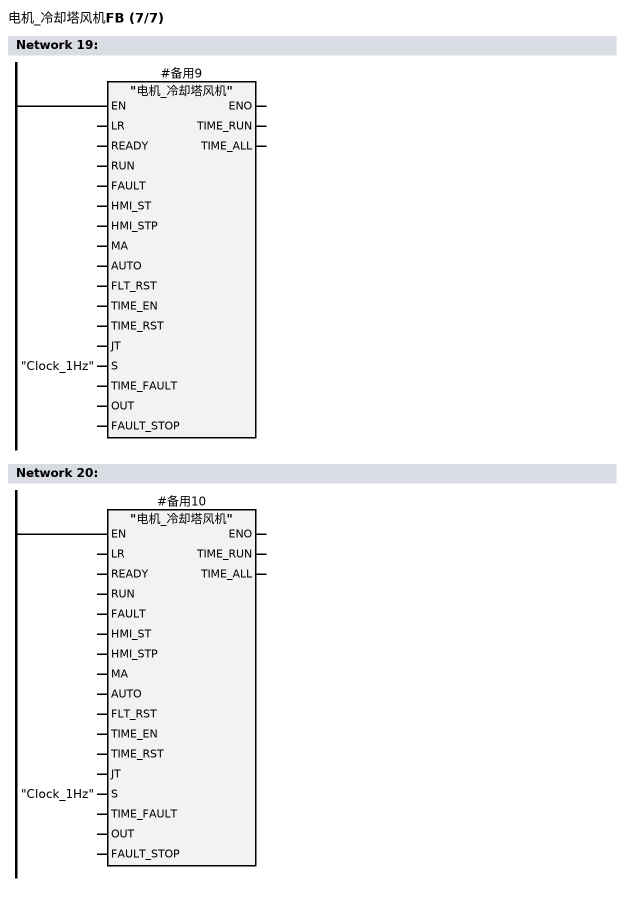
   RUNG wire#powerrail
      #备用9(LR :=, READY :=, RUN :=, FAULT :=, HMI_ST :=, HMI_STP :=, MA :=, AUTO :=, FLT_RST :=, TIME_EN :=, TIME_RST :=, JT :=, S := "Clock_1Hz", TIME_FAULT :=, OUT :=, FAULT_STOP :=, TIME_RUN =>, TIME_ALL =>)
   END_RUNG
   // the same network as SCL:
   #备用9(S := "Clock_1Hz");   // "电机_冷却塔风机"
END_REGION

REGION Network 20
   RUNG wire#powerrail
      #备用10(LR :=, READY :=, RUN :=, FAULT :=, HMI_ST :=, HMI_STP :=, MA :=, AUTO :=, FLT_RST :=, TIME_EN :=, TIME_RST :=, JT :=, S := "Clock_1Hz", TIME_FAULT :=, OUT :=, FAULT_STOP :=, TIME_RUN =>, TIME_ALL =>)
   END_RUNG
   // the same network as SCL:
   #备用10(S := "Clock_1Hz");   // "电机_冷却塔风机"
END_REGION
END_FUNCTION_BLOCK

FUNCTION_BLOCK "阀门_FB"   // FB11, LAD
{ S7_Optimized_Access := 'FALSE' }